(* CODESYS project CodeSys_main.project (continued)
  5ce3da45-db07-42e7-a21c-a00fff4ed8f6|C:\Users\ggb\Documents\#PROJECTS\2016_06_29_Denmark\Visu\RightArrow_Bold.png
  5ce3da45-db07-42e7-a21c-a00fff4ed8f6|C:\Users\ggb\Documents\#PROJECTS\2016_06_29_Denmark\Visu\Parameters_0.png
  5ce3da45-db07-42e7-a21c-a00fff4ed8f6|C:\Users\ggb\Documents\#PROJECTS\2016_06_29_Denmark\Pictures\071-060_Kameraprüfen.jpg
  5ce3da45-db07-42e7-a21c-a00fff4ed8f6|C:\Users\ggb\Documents\#PROJECTS\2016_06_29_Denmark\Visu\Manual_0.png
  5ce3da45-db07-42e7-a21c-a00fff4ed8f6|C:\Users\ggb\Documents\#PROJECTS\2016_06_29_Denmark\Pictures\071-046b_Magazin.jpg
  5ce3da45-db07-42e7-a21c-a00fff4ed8f6|C:\Users\ggb\Documents\#PROJECTS\2016_06_29_Denmark\Pictures\071-050a_Bohren EA.jpg
  5ce3da45-db07-42e7-a21c-a00fff4ed8f6|C:\Users\ggb\Documents\#PROJECTS\2016_06_29_Denmark\Visu\RightArrow_Bold.png
  5ce3da45-db07-42e7-a21c-a00fff4ed8f6|C:\Users\ggb\Documents\#PROJECTS\2016_06_29_Denmark\Visu\Manual_1.png
  5ce3da45-db07-42e7-a21c-a00fff4ed8f6|C:\Users\ggb\Documents\#PROJECTS\2016_06_29_Denmark\Visu\Plus.png
  5ce3da45-db07-42e7-a21c-a00fff4ed8f6|C:\Users\ggb\Documents\#PROJECTS\2016_06_29_Denmark\Visu\LeftArrow_Bold.png
  5ce3da45-db07-42e7-a21c-a00fff4ed8f6|C:\Users\ggb\Documents\#PROJECTS\2016_06_29_Denmark\Visu\German.gif
  5ce3da45-db07-42e7-a21c-a00fff4ed8f6|C:\Users\ggb\Documents\#PROJECTS\2016_06_29_Denmark\Pictures\071-030_Modul Trocknen.jpg
  5ce3da45-db07-42e7-a21c-a00fff4ed8f6|C:\Users\ggb\Documents\#PROJECTS\2016_06_29_Denmark\Visu\CheckBox_1.png
  5ce3da45-db07-42e7-a21c-a00fff4ed8f6|C:\Users\ggb\Documents\#PROJECTS\2016_06_29_Denmark\Visu\Manual_1.png
  5ce3da45-db07-42e7-a21c-a00fff4ed8f6|C:\Users\ggb\Documents\#PROJECTS\2016_06_29_Denmark\Visu\RightArrow.png
  5ce3da45-db07-42e7-a21c-a00fff4ed8f6|C:\Users\ggb\Documents\#PROJECTS\2016_06_29_Denmark\Visu\English.gif
  5ce3da45-db07-42e7-a21c-a00fff4ed8f6|C:\Users\ggb\Documents\#PROJECTS\2016_06_29_Denmark\Pictures\cpFactory_Conveyor.png
  5ce3da45-db07-42e7-a21c-a00fff4ed8f6|C:\Users\ggb\Documents\#PROJECTS\2016_06_29_Denmark\Visu\Parameters_0.png
  5ce3da45-db07-42e7-a21c-a00fff4ed8f6|C:\Users\ggb\Documents\#PROJECTS\2016_06_29_Denmark\Visu\Stopper.jpg
  5ce3da45-db07-42e7-a21c-a00fff4ed8f6|C:\Users\ggb\Documents\#PROJECTS\2016_06_29_Denmark\Visu\RightArrow_Bold.png
  5ce3da45-db07-42e7-a21c-a00fff4ed8f6|C:\Users\ggb\Documents\#PROJECTS\2016_06_29_Denmark\Visu\Home_1.png
  5ce3da45-db07-42e7-a21c-a00fff4ed8f6|C:\Users\ggb\Documents\#PROJECTS\2016_06_29_Denmark\Visu\CheckBox_0.png
  5ce3da45-db07-42e7-a21c-a00fff4ed8f6|C:\Users\ggb\Documents\#PROJECTS\2016_06_29_Denmark\Pictures\071-050a_Bohren EA.jpg
  5ce3da45-db07-42e7-a21c-a00fff4ed8f6|C:\Users\ggb\Documents\#PROJECTS\2016_06_29_Denmark\Visu\German.gif
  5ce3da45-db07-42e7-a21c-a00fff4ed8f6|C:\Users\ggb\Documents\#PROJECTS\2016_06_29_Denmark\Visu\English.gif
  5ce3da45-db07-42e7-a21c-a00fff4ed8f6|C:\Users\ggb\Documents\#PROJECTS\2016_06_29_Denmark\Visu\Plus.png
  5ce3da45-db07-42e7-a21c-a00fff4ed8f6|C:\Users\ggb\Documents\#PROJECTS\2016_06_29_Denmark\Visu\Parameters_1.png
*)

// Data Types/HMI and SCADA/st_WinCC
/////////////////////////////////
/////////////////////////////////
TYPE st_WinCC :
STRUCT
	/// activate Automatic mode
	xAuto: BOOL;
	/// activate Reset mode
	xReset: BOOL;
	/// Stop at cycle end
	xCycleEnd: BOOL;
	/// activate Manual mode
	xManual: BOOL;
	/// activate Teach mode
	xTeach: BOOL;
	/// Quit Error from WinCC
	xQuit: BOOL;
	/// Clear RFID Data (without CarrierID)
	xClrRFID: BOOL;
END_STRUCT
END_TYPE

// Data Types/SAP/sub_structures/st_Par_Req

TYPE st_Par_Req :
STRUCT
	sSfc		: STRING(18);
	sDcGroup	: STRING(12);
	sName1		: STRING(30);
	iValue1		: INT;
	sName2		: STRING(30);
	iValue2		: INT;
	sName3		: STRING(30);
	iValue3		: INT;
	sName4		: STRING(30);
	iValue4		: INT;
	iCamResult	: INT;
END_STRUCT
END_TYPE

// Data Types/Error/st_InteractiveError
//////////////////////////////////////////////
//////////////////////////////////////////////
TYPE st_InteractiveError :
STRUCT
	/// Interactive error is active
	xError: BOOL;
	/// Message ID (ID of the InteractiveErrors textlist row)
	sMessageID: STRING;
	/// The actual state of the stopper
	uiState: UINT;
	/// The state of stopper after pushing the Ignore button
	uiIgnoreState: UINT;
	/// The state of stopper after pushing the Abort button
	uiAbortState: UINT;
	/// Repeat button was pushed
	xBtnRepeat: BOOL;
	/// Ignore button was pushed
	xBtnIgnore: BOOL;
	/// Abort button was pushed
	xBtnAbort: BOOL;
	// Reject order button was pushed
	xBtnRejectOrder: BOOL;
END_STRUCT
END_TYPE

// Data Types/HMI and SCADA/CDPX/st_StopperSensorSignals
TYPE st_StopperSensorSignals :
STRUCT
	xInductive_1		: BOOL;
	xInductive_2		: BOOL;
	xInductive_3		: BOOL;
	xInductive_4		: BOOL;
	xStpDownSensor		: BOOL;
	xStpDownOutpu		: BOOL;
	sInductive_1		: STRING(5);
	sInductive_2		: STRING(5);
	sInductive_3		: STRING(5);
	sInductive_4		: STRING(5);
	sStpDownSensor		: STRING(5);
	sStpDownOutpu		: STRING(5);
	sRfid				: STRING(5);
	xTagPresent			: BOOL;
	xReady				: BOOL;
	xBusy				: BOOL;
	xError				: BOOL;
	xTimeOut			: BOOL;		
END_STRUCT
END_TYPE

// Data Types/HMI and SCADA/st_ManualWorkplace
TYPE st_ManualWorkplace :
STRUCT
	sURL				: STRING;
	xManualJob			: BOOL;
	xManualJobStarted	: BOOL;
	xManualJobFinished	: BOOL;
	xManualJobCanceled	: BOOL;
END_STRUCT
END_TYPE

// Data Types/HMI and SCADA/CDPX/st_InterctiveErrors
TYPE st_InterctiveErrors :
STRUCT
	xIntDefault		: BOOL;
	xIntMES			: BOOL;
	xIntSAP			: BOOL;
	xIntApp			: BOOL;
	xIntMan			: BOOL;
	xIntKuka		: BOOL;
	
	sURL			: STRING;
	uiIntMsgID		: UINT;
	uiIntState		: UINT;
	uiIntIgnore		: UINT;
	uiIntAbort		: UINT;
	uiSapOp			: UDINT;
	uiSapPos		: UDINT;
	sSapError		: STRING;
	udiSapSfc		: UDINT;	
END_STRUCT
END_TYPE

// Data Types/HMI and SCADA/CDPX/st_Errors
TYPE st_Errors :
STRUCT
	xError			: BOOL;
	uiLevel			: UINT;
	uiMsgNum		: UINT;
	sErrorID		: STRING[4);
	sDateTime		: STRING;
END_STRUCT
END_TYPE

// Data Types/Error/st_RobotError
TYPE st_RobotError :
STRUCT
	/// Interactive error is active
	xError: BOOL;
	/// Message ID (ID of the InteractiveErrors textlist row)
	sMessageID: STRING;
	/// The state of stopper after pushing the Retry button
	uiRetryState: UINT;
	/// The state of stopper after pushing the Exit button
	uiExitState: UINT;
	/// Retry button was pushed
	xBtnRetry: BOOL;
	/// Exit button was pushed
	xBtnExit: BOOL;
END_STRUCT
END_TYPE

// Data Types/Application/st_AppControl
TYPE st_AppControl :
STRUCT
	xStart		: BOOL;
	xReset		: BOOL;
	xStop		: BOOL;
	uiOpNo		: UINT;
	auiPar		: ARRAY [0..3] OF UINT;
	udiONo		: UDINT;
	uiOPos		: UINT;
END_STRUCT
END_TYPE

// Data Types/HMI and SCADA/CDPX/st_ConveyorSignals
TYPE st_ConveyorSignals :
STRUCT
	xConvMovingLeft		: BOOL;
	xConvMovingRight	: BOOL;
	xConvMovingSlow		: BOOL;
	
	sConvLeft			: STRING(5);
	sConvRight			: STRING(5);
	sConvSlow			: STRING(5);	
END_STRUCT
END_TYPE

// Data Types/Error/u_Error
////////////////////////////////////////////////////////////////////////////////////////
/////////////////////////////////////////////////////////////////////////////////////////
TYPE u_Error :

UNION
	/// Long Word (64 bit) for error bits
	lwError: LWORD;
	/// 4 times Word for WinCC visualization
	stErrorWords: st_ErrorWords;
END_UNION

END_TYPE

// Data Types/Error/st_Error
///////////////////////////////////
///////////////////////////////////
TYPE st_Error :
STRUCT
	/// Union to store Level 0 errors in LWORD and 4xWORD for WinCC
	uL0: u_Error;
	/// Union to store Level 1 errors in LWORD and 4xWORD for WinCC
	uL1: u_Error;
	/// Union to store Level 2 errors in LWORD and 4xWORD for WinCC	
	uL2: u_Error;
	/// Error flags
	xSF0: BOOL;
	/// summary error flag Level 1
	xSF1: BOOL;
	/// summary error flag Level 2
	xSF2: BOOL;
	/// global error flag (SF0 or SF1)
	xSF: BOOL;
	/// extended (100ms) global error flag
	xSF_ext: BOOL;
	/// confirm error
	xQuit: BOOL;
END_STRUCT
END_TYPE

// Data Types/SAP/sub_structures/st_Start_Req

TYPE st_Start_Req :
STRUCT
	sSfc	: STRING(18);
	sItem	: STRING(18);
END_STRUCT
END_TYPE

// Data Types/SAP/st_CompleteSfc

TYPE st_CompleteSfc :
STRUCT
	Req		: st_Comp_Req;
	Res		: st_Comp_Res;
	Com		: st_Com;
END_STRUCT
END_TYPE

// Data Types/HMI and SCADA/st_ButtonState
TYPE st_ButtonState :
STRUCT
	xPressed	: BOOL;
	xActive		: BOOL;
	xDisabled	: BOOL;
END_STRUCT
END_TYPE

// Data Types/SAP/st_ParametricData

TYPE st_ParametricData :
STRUCT
	Req		: st_Par_Req;
	Com		: st_Com;
END_STRUCT
END_TYPE

// Data Types/Application/st_AppSettings
TYPE st_AppSettings :
STRUCT
	xActive			: BOOL := TRUE;
	xStopBelt		: BOOL;
	xCarrierInit	: BOOL;
	uiCarrierInitNum: UINT := 1;
END_STRUCT
END_TYPE

// Data Types/HMI and SCADA/CDPX/st_AppButtonControl
TYPE st_AppButtonControl :
STRUCT
	xButton		: BOOL;
	sButton		: STRING(16);	
END_STRUCT
END_TYPE

// Data Types/SAP/sub_structures/st_Com

TYPE st_Com :
STRUCT
	iTrigger		: INT;
	iResponse		: INT;
	bError			: BIT;
	sError			: STRING(128);
END_STRUCT
END_TYPE

// Data Types/Application/st_AppState
TYPE st_AppState :
STRUCT
	xReady					: BOOL;
	xError					: BOOL;
	xInitPos				: BOOL;
	uiReturnCode			: UINT;
END_STRUCT
END_TYPE

// Data Types/HMI and SCADA/CDPX/st_StopperButtonState
TYPE st_StopperButtonState :
STRUCT
	xInit		: BOOL;
	xRead		: BOOL;
	xWrite		: BOOL;
	xDeleteData	: BOOL;
	xStpMveDown	: BOOL;
	xStpMveUp	: BOOL;
END_STRUCT
END_TYPE

// Data Types/Error/st_ErrorWords
/////////////////////////
/////////////////////////
TYPE st_ErrorWords :
STRUCT
	wErrorWord0: WORD;
	wErrorWord1: WORD;
	wErrorWord2: WORD;
	wErrorWord3: WORD;
END_STRUCT
END_TYPE

// Data Types/SAP/sub_structures/st_Start_Res

TYPE st_Start_Res :
STRUCT
	sDcGroup	: STRING(12);
	sName1		: STRING(30);
	iValue1		: INT;
	sName2		: STRING(30);
	iValue2		: INT;
	sName3		: STRING(30);
	iValue3		: INT;
	sName4		: STRING(30);
	iValue4		: INT;
	sItem		: STRING(18);
	sItemRev	: STRING(3);
	sSfc		: STRING(10);	
END_STRUCT
END_TYPE

// Data Types/HMI and SCADA/CDPX/st_CdpxButtonState
TYPE st_CdpxButtonState :
STRUCT
	xClearError		: BOOL;
	xOperationMode	: BOOL;
	xOverview     	: BOOL;
	xUser         	: BOOL;
	xHome         	: BOOL;
	xSetupMode    	: BOOL;
	xParameter    	: BOOL;
	xSystem       	: BOOL;
	xApp_1        	: BOOL;
	xApp_2        	: BOOL;
	xStp_1        	: BOOL;
	xStp_2        	: BOOL;
	xBelt         	: BOOL;
	xApp          	: BOOL;
	xTrans_1      	: BOOL;
	xTrans_2      	: BOOL;
	xSwLanguage		: BOOL;
	xCloseDialog	: BOOL;
END_STRUCT
END_TYPE

// Data Types/SAP/ManualWork/st_MesRcvData_ManualWork
TYPE st_MesRcvData_ManualWork :
STRUCT
	stHeader		: dc_ecp.st_MES4_QueryHeader;
	sOderDes		: STRING[60];
	sPartDes		: STRING[20];
END_STRUCT
END_TYPE

// Data Types/Application/st_AppInfo
TYPE st_AppInfo :
STRUCT
	auiOperations			: ARRAY [0..15] OF UINT;
	byNumberOfOperations	: BYTE;
END_STRUCT
END_TYPE

// Data Types/SAP/sub_structures/st_Comp_Req

TYPE st_Comp_Req :
STRUCT
	sSfc	: STRING(18);
END_STRUCT
END_TYPE

// Data Types/HMI and SCADA/CDPX/st_AppSensors
TYPE st_AppSensors :
STRUCT
	xSensor		: BOOL;
	sSensor		: STRING(16);
END_STRUCT
END_TYPE

// Data Types/SAP/sub_structures/st_Comp_Res

TYPE st_Comp_Res :
STRUCT
	sOp		: STRING(4);
	sOpRev	: STRING(3);
END_STRUCT
END_TYPE

// Data Types/st_GetShuntId
TYPE st_GetShuntId :
STRUCT
	uiSourceId			: UINT;
	uiSourcePosition	: UINT;
	uiTargetId			: UINT;
	uiTargetPosition	: UINT;
END_STRUCT
END_TYPE

// Data Types/Error/st_ErrorEvent
///////////////////////////////////
///////////////////////////////////
TYPE st_ErrorEvent :
STRUCT
	/// Error ID (ID of the Errors textlist row)
	sErrorID: STRING := 'No error';
	/// Text message (It does not contains anyting, it is only to show an additional column in the visualization)
	sErrorText: STRING;
	/// String of the date and time
	sDateTime: STRING;
END_STRUCT
END_TYPE

// Data Types/HMI and SCADA/st_TransitionData
TYPE st_TransitionData :
STRUCT
	uiCondIn	: UINT;
	uiPar1		: UINT;
	uiPar2		: UINT;
	uiPar3		: UINT;
	uiPar4		: UINT;
	xAppEn		: BOOL;
	uiCondOut	: UINT;
	uiCondAbort	: UINT;
	byStopper	: BYTE;
END_STRUCT
END_TYPE

// Data Types/SAP/st_StartSfc

TYPE st_StartSfc :
STRUCT
	Req	: st_Start_Req;
	Res	: st_Start_Res;
	Com	: st_Com;
END_STRUCT
END_TYPE

// Data Types/HMI and SCADA/CDPX/st_ConveyorButtonState
TYPE st_ConveyorButtonState :
STRUCT
	xConvLeft		: BOOL;
	xConvRight		: BOOL;
	xConvSlow		: BOOL;
END_STRUCT
END_TYPE

// Global Variables/fromCDPX
{attribute 'qualified_only'}
VAR_GLOBAL
	uiMode									: UINT;
	uiDummy									: UINT;
	stCdpxButtonState						: st_CdpxButtonState;
	
	
	stHome_OperationMode_Reset		 		: st_ButtonState;
	stHome_OperationMode_Automatic		 	: st_ButtonState;
	stHome_OperationMode_Setup 				: st_ButtonState;
	stHome_OperationMode_CycleEnd 			: st_ButtonState;
	
	stSetupMode_Stopper1_Init		 		: st_ButtonState;
	stSetupMode_Stopper1_Read			 	: st_ButtonState;
	stSetupMode_Stopper1_Write 				: st_ButtonState;
	stSetupMode_Stopper1_DeleteData 		: st_ButtonState;

	stSetupMode_Stopper2_Init		 		: st_ButtonState;
	stSetupMode_Stopper2_Read			 	: st_ButtonState;
	stSetupMode_Stopper2_Write 				: st_ButtonState;
	stSetupMode_Stopper2_DeleteData 		: st_ButtonState;
	
	stInteractiveMessage_Repeat 			: st_ButtonState;
	stInteractiveMessage_Ignore	 			: st_ButtonState;
	stInteractiveMessage_Abort				: st_ButtonState;	
	stInteractiveMessage_RejectOrder		: st_ButtonState;	
	
	stManualWorkplace						: st_ManualWorkplace;
	stRobotError							: st_RobotError;	
	astStopperButton						: ARRAY [0..1] OF st_StopperButtonState;
	astAppSetting							: ARRAY [0..1] OF st_AppSettings;
	astAppButtonControl						: ARRAY [0..15] OF st_AppButtonControl;
	astTransitionTable_1					: ARRAY [0..10] OF st_TransitionData;
	astTransitionTable_2					: ARRAY [0..10] OF st_TransitionData;	
	astConveyorButtonState					: ARRAY [0..2] OF st_ConveyorButtonState; 
END_VAR

// APP_FILLING/Application/IO
//{attribute 'qualified_only'} - removed to access variables without "DigitalIO." 
VAR_GLOBAL
	// Application Type Identifier
	xAppID AT %QX0.7: BOOL := TRUE;
	// Push Piston forward
	xPistonOn AT %QX0.0: BOOL := FALSE;
	// Turns pump on
	xPumpOn AT %QX0.2: BOOL := FALSE;
	// Indicates if the app is powered on or off
	xIsOn AT %QX0.6: BOOL := TRUE;
	// Indicates which module (09 or 08) the app is mounted on
	xModuleID AT %IX0.7: BOOL;
END_VAR

// Global Variables/Standards
VAR_GLOBAL
	/// First-Cycle-Flag
	xFirstCycle: BOOL := TRUE;
	/// Initialization flag
	xInit: BOOL;
	/// Station is in Initial Position
	xInitPos: BOOL;
	/// Startup like warmstart
	xSoftReset: BOOL;
	/// Application program is idle	
	xAppIdle: BOOL;
	/// Application program is busy
	xAppBusy: BOOL;
	/// Automatic Mode is active
	xAuto: BOOL;
	/// Automatic Start is enable
	xAutoEn: BOOL;
	/// Reset Mode is active
	xReset: BOOL;
	/// Reset Start is enable
	xResetEn: BOOL;
	/// Reset sequence is finished
	xResetRdy: BOOL;
	/// Manual Mode is active
	xManual: BOOL;
	/// Manual Start is enable
	xManualEn: BOOL;
	/// Teach Mode is active	
	xTeach: BOOL;
	/// Teach Start is enable
	xTeachEn: BOOL;
	/// Stop at cycle end is active	
	xCycleEnd: BOOL;
	/// Stop at cycle end is enable
	xCycleEndEn: BOOL;
	/// Reset Automatic Start flag
	xAutoReset: BOOL := FALSE;
	/// Stopper ST1 in idle state          		
	xSt1_Idle: BOOL;
	/// Stopper ST2 in idle state          		
	xSt2_Idle: BOOL;
	/// Stopper ST2 in idle state          		
	xSt3_Idle: BOOL;
	/// Resource is busy
	xBusy: BOOL;
	/// MES mode is active
	xMES: BOOL;
	/// SAP mode is active
	xSAP: BOOL;
	/// Struct with 64 Error Flags
	stError: st_Error;
	/// Structure with WinCC variables     
	stWinCC: st_WinCC;
	/// Structure with HMI variables
	stHMI: st_WinCC;
	//Semaphore for gate
	xSema : BOOL;
	// Semaphore for shunt
	xSemaShunt	: BOOL;
END_VAR

// Global Variables/toCDPX
{attribute 'qualified_only'}
VAR_GLOBAL
	sModule						: STRING(32);
	byOpMode					: BYTE;
	byScreenTitle				: BYTE;
	xManual						: BOOL;
	xAuto						: BOOL;
	xSAP						: BOOL;
	xMES						: BOOL;
	xDefault					: BOOL;
	auiCarrierInitNum			: ARRAY [0..1] OF UINT;
	uiNumOfApplications			: UINT;
	uiNumOfStoppers				: UINT;
	uiNumOfBelts				: UINT;
	auiCondIn					: ARRAY [0..1] OF UINT;
	auiCondOut					: ARRAY [0..1] OF UINT;
	sTime						: STRING;
	sDate						: STRING;
	stInteractiveErrors			: st_InterctiveErrors;
	astErrors					: ARRAY [1..20] OF st_Errors;
	astRfidData					: ARRAY [0..1] OF dc_ecp.st_CPF_VisuData;
	astSensorSignals			: ARRAY [0..1] OF st_StopperSensorSignals;
	astConveyorSignals			: ARRAY [0..2] OF st_ConveyorSignals;
	astAppState					: ARRAY [0..1] OF st_AppState;
	astAppControl				: ARRAY [0..1] OF st_AppControl;	
	astAppSensors				: ARRAY [0..31] OF st_AppSensors;
	auiValues					: ARRAY [0..31] OF UINT;	
	astAppControlONo: UDINT := 0;
END_VAR

// Global Variables/SAP
{attribute 'qualified_only'}
VAR_GLOBAL
	Start			: st_StartSfc;
	Par				: st_ParametricData;
	Comp			: st_CompleteSfc;
END_VAR

// Global Variables/SAPInit
{attribute 'qualified_only'}
VAR_GLOBAL
	Start			: st_StartSfc;
	Par				: st_ParametricData;
	Comp			: st_CompleteSfc;
END_VAR

// Global Variables/SAPHMI
{attribute 'qualified_only'}
VAR_GLOBAL
	uiOp		: UDINT;
	uiPos		: UDINT;
	sError		: STRING;
	udiSfc		: UDINT;	
END_VAR

// MODULE_PLC09/Application/Variables/IO
VAR_GLOBAL
	

	///////////////////////////
	// Inputs
	///////////////////////////
	
	xBG20		AT %IX1.0	: BOOL;	// Stopper released
	xBG21		AT %IX1.1	: BOOL;	// Carrier available
	xBG22		AT %IX1.2	: BOOL;	// Carrier ID bit 0
	xBG23		AT %IX1.3	: BOOL;	// Carrier ID bit 1
	xBG24		AT %IX1.4	: BOOL;	// Carrier ID bit 2
	xEmg		AT %IX0.0	: BOOL;	// Emergency stop
	
	///////////////////////////
	// Outputs
	///////////////////////////	
	
	xMB20		AT %QX1.0	: BOOL;	// Release stopper
	xQA1_LEFT	AT %QX0.5	: BOOL;	// Conveyor to the left
	xQA1_RIGHT	AT %QX0.4	: BOOL;	// Conveyor to the right
	xQA1_SLOW	AT %QX0.6	: BOOL;	// Conveyor Slow
	xQA1_STOP	AT %QX0.7	: BOOL;	// Conveyor Stop
	// Application Identifier
	xAPP_ID AT %IX0.1: BOOL;
	
	
	
	
	// Application power status
	xAppIsOn AT %IX0.2: BOOL;
	// Module Identifier Bit
	xModuleID AT %QX0.0: BOOL := FALSE;
END_VAR

// MODULE_PLC09/Application/Variables/NVL_PLC09_REC_FILLING
//This gobal variable list is received via the network.
//Sender: NVL_FILLING_SEND [APP_FILLING: PLC Logic: Application]
//Protocol: UDP

VAR_GLOBAL
	isDone: BOOL := FALSE;
	isOn: BOOL := FALSE;
END_VAR

// MODULE_PLC09/Application/Variables/NVL_PLC09_SEND
VAR_GLOBAL
	Ready: BOOL := FALSE;
END_VAR

// MODULE_PLC08/Application/Variables/IO
VAR_GLOBAL
	

	///////////////////////////
	// Inputs
	///////////////////////////
	
	xBG20		AT %IX1.0	: BOOL;	// Stopper released
	xBG21		AT %IX1.1	: BOOL;	// Carrier available
	xBG22		AT %IX1.2	: BOOL;	// Carrier ID bit 0
	xBG23		AT %IX1.3	: BOOL;	// Carrier ID bit 1
	xBG24		AT %IX1.4	: BOOL;	// Carrier ID bit 2
	xEmg		AT %IX0.0	: BOOL;	// Emergency stop
	
	///////////////////////////
	// Outputs
	///////////////////////////	
	
	xMB20		AT %QX1.0	: BOOL;	// Release stopper
	xQA1_LEFT	AT %QX0.5	: BOOL;	// Conveyor to the left
	xQA1_RIGHT	AT %QX0.4	: BOOL;	// Conveyor to the right
	xQA1_SLOW	AT %QX0.6	: BOOL;	// Conveyor Slow
	xQA1_STOP	AT %QX0.7	: BOOL;	// Conveyor Stop
	// Application Identifier
	xAPP_ID AT %IX0.1: BOOL;
	
	
	// Application power status
	xAppIsOn AT %IX0.2: BOOL;
	// Module Identifier Bit
	xModuleID AT %QX0.0: BOOL := TRUE;
END_VAR

// MODULE_PLC08/Application/Variables/NVL_PLC08_SEND
VAR_GLOBAL
	Ready: BOOL := FALSE;
END_VAR

// APP_FILLING/Application/NVL_FILLING_SEND
VAR_GLOBAL
	isDone: BOOL := FALSE;
	isOn: BOOL := FALSE;
END_VAR

// APP_FILLING/Application/NVL_FILLING_REC_09
//This gobal variable list is received via the network.
//Sender: NVL_PLC09_SEND [MODULE_PLC09: PLC Logic: Application]
//Protocol: UDP

VAR_GLOBAL
	Ready: BOOL := FALSE;
END_VAR

// APP_STOPPERING/Application/IO
//{attribute 'qualified_only'} - removed to access variables without "DigitalIO." 
VAR_GLOBAL
	// Application Type Identifier
	xAppID AT %QX0.7: BOOL := FALSE;
	// Push Piston forward
	xPistonOn AT %QX0.0: BOOL := FALSE;
	// Pushes stoppering down to the containers
	xStopperingOn AT %QX0.2: BOOL := FALSE;
	// Indicates if the app is powered on or off
	xIsOn AT %QX0.6: BOOL := TRUE;
	// Indicates which module (09 or 08) the app is mounted on
	xModuleID AT %IX0.7: BOOL;
END_VAR

// APP_STOPPERING/Application/NVL_STOPPERING_SEND
VAR_GLOBAL
	isDone: BOOL := FALSE;
END_VAR

// APP_STOPPERING/Application/NVL_STOPPERING_REC_08
//This gobal variable list is received via the network.
//Sender: NVL_PLC08_SEND [MODULE_PLC08: PLC Logic: Application]
//Protocol: UDP

VAR_GLOBAL
	Ready: BOOL := FALSE;
END_VAR

// MODULE_PLC08/Application/Variables/NVL_PLC08_REC_STOPPERING
//This gobal variable list is received via the network.
//Sender: NVL_STOPPERING_SEND [APP_STOPPERING: PLC Logic: Application]
//Protocol: UDP

VAR_GLOBAL
	isDone: BOOL := FALSE;
END_VAR

// MODULE_PLC08/Application/Variables/NVL_PLC08_REC_FILLING
//This gobal variable list is received via the network.
//Sender: NVL_FILLING_SEND [APP_FILLING: PLC Logic: Application]
//Protocol: UDP

VAR_GLOBAL
	isDone: BOOL := FALSE;
	isOn: BOOL := FALSE;
END_VAR

// APP_STOPPERING/Application/NVL_STOPPERING_REC_09
//This gobal variable list is received via the network.
//Sender: NVL_PLC09_SEND [MODULE_PLC09: PLC Logic: Application]
//Protocol: UDP

VAR_GLOBAL
	Ready: BOOL := FALSE;
END_VAR

// APP_FILLING/Application/NVL_FILLING_REC_08
//This gobal variable list is received via the network.
//Sender: NVL_PLC08_SEND [MODULE_PLC08: PLC Logic: Application]
//Protocol: UDP

VAR_GLOBAL
	Ready: BOOL := FALSE;
END_VAR

// MODULE_PLC09/Application/Variables/NVL_PLC09_REC_STOPPERING
//This gobal variable list is received via the network.
//Sender: NVL_STOPPERING_SEND [APP_STOPPERING: PLC Logic: Application]
//Protocol: UDP

VAR_GLOBAL
	isDone: BOOL := FALSE;
END_VAR

// MODULE_PLC09/Application/Programs/MODULE_PLC09_MAIN
PROGRAM  MODULE_PLC09_MAIN
VAR
	state: UINT := 0;
	PLCid: STRING;
	RFID: dc_ecp.Dtm425;
	RfidData: dc_ecp.st_CPF_RfidData;
	ConveyorRight: BOOL;
	CarrierID: UINT := 0;
	TIMER: TON;
	WaitTime: TIME;
	AppType: STRING;
	PistonState: STRING := 'retracted';
	ServerCommand: STRING := 'wait';
	AppState: STRING := 'waiting';
	CarrierIdString: STRING := '0';
END_VAR

CASE state OF
	
	0: // init
	IO.xMB20 := FALSE; // raise stoppper
	RFID.ClearError();
	PLCid := 'STPLC_09';
	state := 5;
	
	5: // identify
	AppState := 'N/A';
	IF IO.xAppIsOn THEN
		IF IO.xAPP_ID THEN
			AppType := 'filling';
		ELSE
			AppType := 'stoppering';
		END_IF
		state:=10;
	END_IF
	
	10: // wait for RFID to clear
	AppState := 'starting';
	IF RFID.xReady THEN
		RFID.Connect(32, 0, 1);
		state:=20;
	END_IF
	
	20: // wait for RFID be ready then move conveyor
	//CarrierID := 0;
	IF RFID.xReady AND IO.xAppIsOn THEN
		AppState := 'ready';
		IF ServerCommand = 'begin' THEN
			AppState := 'waiting';
			IO.xMB20 := TRUE;
			IO.xQA1_RIGHT := TRUE; // Move conveyor right
			state:=30;
		END_IF
	ELSE
		AppState := 'N/A';
	END_IF
	
	30: // wait for carrier to be available
	IF IO.xBG21 THEN
		IO.xQA1_RIGHT := FALSE; // stop conveyor
		IO.xMB20 := FALSE; // lower stoppper
		state:=40;
	END_IF
	
	
	40: // wait for RFID to read then send
	IF RFID.xReady THEN
		RFID.ReadTag(uiStartAddress := 0, uiDataLength := SIZEOF(RfidData), ADR(RfidData));
		state := 42;
	END_IF
	
	42:
	IF RFID.xReady THEN
		CarrierID := dc_ecp.SwapWord(RfidData.uiCarrierID); // swap bit order
		
		IF CarrierID > 0 THEN
			AppState := 'ready';
			state := 45;
		ELSE
			AppState := 'waiting';
		END_IF
	END_IF
	
	45: // wait for server to tell if pass or go
	IF ServerCommand = 'valid' THEN
		IF AppType = 'filling' THEN
			AppState := 'filling';
			state := 46;
		ELSIF AppType = 'stoppering' THEN
			AppState := 'stoppering';
			state := 46;
		END_IF
	ELSIF ServerCommand = 'pass' THEN
		AppState := 'passing';
		state := 100;
	END_IF
	
	46:
	NVL_PLC09_SEND.Ready := TRUE;
	WaitTime := STRING_TO_TIME('T#500ms');
	TIMER(IN := TRUE, PT := WaitTime);
	IF TIMER.Q = TRUE THEN 
		TIMER(IN := FALSE);
		NVL_PLC09_SEND.Ready := FALSE;
		state := 50;
	END_IF
	
	
	50: // wait for task to complete, then report back
	IF AppType = 'stoppering' THEN
		IF NVL_PLC09_REC_STOPPERING.isDone THEN
			AppState := 'done';
			state := 55;
		END_IF
	ELSIF AppType = 'filling' THEN
		IF NVL_PLC09_REC_FILLING.isDone THEN
			AppState := 'done';
			state := 55;
		END_IF
	END_IF
	
	55: // wait for server to tell it to move on
	IF ServerCommand = 'transfer' THEN
		state := 100;
	END_IF
	

	
	100: // pass move conveyor again, give 1 sec breathing room
	IO.xMB20 := TRUE; // release stopper
	IF IO.xBG20 THEN // checks if stopper has been released
		IO.xQA1_RIGHT := TRUE; // move conveyor right
		WaitTime := STRING_TO_TIME('T#2000ms');
		timer(IN:=TRUE,PT:=WaitTime);
		state := 105;
	END_IF
	
	105: // wait for timer then restart
	IF timer.Q = TRUE THEN
		timer(IN:=FALSE);
		IF ServerCommand = 'pass' THEN
			AppState := 'passed';
		ELSIF ServerCommand = 'transfer' THEN
			AppState := 'done';
		END_IF
		state := 30;
		CarrierID := 0;
		ServerCommand := 'begin';
	END_IF
	
	
	
END_CASE
RFID();
timer();

END_PROGRAM

// APP_FILLING/Application/APP_FILLING_MAIN
PROGRAM APP_FILLING_MAIN
VAR
	state: UINT := 0;
	APPid: STRING;
	TIMER: TON;
	WaitTime: TIME;
	ModuleID: STRING;
END_VAR

CASE state OF
	
	0: // init
	APPid := 'APP_FILLINGs';
	IO.xPistonOn := FALSE;
	IO.xPumpOn := FALSE;
	IO.xIsOn := TRUE;
	IO.xAppID := TRUE;
	NVL_FILLING_SEND.isOn := TRUE;
	state := 10;
	
	10: //  Read Module id
	IF IO.xModuleID = TRUE THEN
		ModuleID := '08';
	ELSIF IO.xModuleID = FALSE THEN
		ModuleID := '09';
	END_IF
	state := 15;
	
	15: // wait for module to be ready
	IF ModuleID = '08' THEN
		IF NVL_FILLING_REC_08.Ready THEN
			NVL_FILLING_SEND.isDone := FALSE;
			state := 20;
		END_IF
	ELSIF ModuleID = '09' THEN
		IF NVL_FILLING_REC_09.Ready THEN
			NVL_FILLING_SEND.isDone := FALSE;
			state := 20;
		END_IF
	END_IF
	
	20: // Push piston forward and wait 5 sec
	IO.xPistonOn := TRUE;
	WaitTime := STRING_TO_TIME ('T#500ms'); // Converts text string to time value --> WaitTime is then 5 sec
	TIMER(IN := TRUE, PT := WaitTime); // Activates the timer and the timers preset time --> The time where the piston is active
	IF Timer.Q = TRUE THEN 
		TIMER(IN := FALSE);
		state := 25;
	END_IF
	
	25: // activate pump for 200ms
	//IO.PistonOn := FALSE;
	IO.xPumpOn := TRUE;
	WaitTime := STRING_TO_TIME ('T#200ms'); // Converts text string to time value --> WaitTime is then 5 sec
	TIMER(IN := TRUE, PT := WaitTime); // Activates the timer and the timers preset time --> The time where the piston is active
	IF Timer.Q = TRUE THEN 
		TIMER(IN := FALSE);
		IO.xPumpOn := FALSE;
		state := 30;
	END_IF
	
	30: // Push piston backwards
	WaitTime := STRING_TO_TIME('T#500ms');
	TIMER(IN := TRUE, PT := WaitTime);
	IF TIMER.Q = TRUE THEN 
		TIMER(IN := FALSE);
		IO.xPistonOn := FALSE;
		state := 40;
	END_IF
	
	40: // Restart conveyor belts
	NVL_FILLING_SEND.isDone := TRUE;
	WaitTime := STRING_TO_TIME('T#1000ms');
	TIMER(IN := TRUE, PT := WaitTime);
	IF TIMER.Q = TRUE THEN 
		TIMER(IN := FALSE);
		state := 15;
	END_IF
	
END_CASE

TIMER();

END_PROGRAM

// MODULE_PLC08/Application/Programs/MODULE_PLC08_MAIN
PROGRAM  MODULE_PLC08_MAIN
VAR
	state: UINT := 0;
	PLCid: STRING;
	RFID: dc_ecp.Dtm425;
	RfidData: dc_ecp.st_CPF_RfidData;
	ConveyorRight: BOOL;
	CarrierID: UINT := 0;
	TIMER: TON;
	WaitTime: TIME;
	AppType: STRING;
	PistonState: STRING := 'retracted';
	ServerCommand: STRING := 'wait';
	AppState: STRING := 'waiting';
END_VAR

CASE state OF
	
	0: // init
	IO.xMB20 := FALSE; // raise stoppper
	RFID.ClearError();
	PLCid := 'STPLC_08';
	state := 5;
	
	5: // identify
	AppState := 'N/A';
	IF IO.xAppIsOn THEN
		IF IO.xAPP_ID THEN
			AppType := 'filling';
		ELSE
			AppType := 'stoppering';
		END_IF
		state:=10;
	END_IF
	
	10: // wait for RFID to clear
	AppState := 'starting';
	IF RFID.xReady THEN
		RFID.Connect(32, 0, 1);
		state:=20;
	END_IF
	
	20: // wait for RFID be ready then move conveyor
	//CarrierID := 0;
	IF RFID.xReady AND IO.xAppIsOn THEN
		AppState := 'ready';
		IF ServerCommand = 'begin' THEN
			AppState := 'waiting';
			IO.xMB20 := TRUE;
			IO.xQA1_RIGHT := TRUE; // Move conveyor right
			state:=30;
		END_IF
	ELSE
		AppState := 'N/A';
	END_IF
	
	30: // wait for carrier to be available
	IF IO.xBG21 THEN
		IO.xQA1_RIGHT := FALSE; // stop conveyor
		IO.xMB20 := FALSE; // lower stoppper
		state:=40;
	END_IF
	
	
	40: // wait for RFID to read then send
	IF RFID.xReady THEN
		RFID.ReadTag(uiStartAddress := 0, uiDataLength := SIZEOF(RfidData), ADR(RfidData));
		state := 42;
	END_IF
	
	42:
	IF RFID.xReady THEN
		CarrierID := dc_ecp.SwapWord(RfidData.uiCarrierID); // swap bit order
		
		IF CarrierID > 0 THEN
			AppState := 'ready';
			state := 45;
		ELSE
			AppState := 'waiting';
		END_IF
	END_IF
	
	45: // wait for server to tell if pass or go
	IF ServerCommand = 'valid' THEN
		IF AppType = 'filling' THEN
			AppState := 'filling';
			state := 46;
		ELSIF AppType = 'stoppering' THEN
			AppState := 'stoppering';
			state := 46;
		END_IF
	ELSIF ServerCommand = 'pass' THEN
		AppState := 'passing';
		state := 100;
	END_IF
	
	46: // tell app to start then wait
	NVL_PLC08_SEND.Ready := TRUE;
	WaitTime := STRING_TO_TIME('T#500ms');
	TIMER(IN := TRUE, PT := WaitTime);
	IF TIMER.Q = TRUE THEN 
		TIMER(IN := FALSE);
		NVL_PLC08_SEND.Ready := FALSE;
		state := 50;
	END_IF
	
	
	50: // wait for task to complete, then report back
	IF AppType = 'stoppering' THEN
		IF NVL_PLC08_REC_STOPPERING.isDone THEN
			AppState := 'done';
			state := 55;
		END_IF
	ELSIF AppType = 'filling' THEN
		IF NVL_PLC08_REC_FILLING.isDone THEN
			AppState := 'done';
			state := 55;
		END_IF
	END_IF
	
	55: // wait for server to tell it to move on
	IF ServerCommand = 'transfer' THEN
		state := 100;
	END_IF
	

	
	100: // pass move conveyor again, give 1 sec breathing room
	IO.xMB20 := TRUE; // release stopper
	IF IO.xBG20 THEN // checks if stopper has been released
		IO.xQA1_RIGHT := TRUE; // move conveyor right
		WaitTime := STRING_TO_TIME('T#2000ms');
		timer(IN:=TRUE,PT:=WaitTime);
		state := 105;
	END_IF
	
	105: // wait for timer then restart
	IF timer.Q = TRUE THEN
		timer(IN:=FALSE);
		IF ServerCommand = 'pass' THEN
			AppState := 'passed';
		ELSIF ServerCommand = 'transfer' THEN
			AppState := 'done';
		END_IF
		state := 20;
		CarrierID := 0;
		ServerCommand := 'begin';
	END_IF
	
	
	
END_CASE
RFID();
timer();

END_PROGRAM

// APP_STOPPERING/Application/APP_STOPPERING_MAIN
PROGRAM APP_STOPPERING_MAIN
VAR
	state: UINT := 0;
	APPid: STRING;
	TIMER: TON;
	WaitTime: TIME;
	ModuleID: STRING;
END_VAR

CASE state OF
	
	0: // init
	APPid := 'APP_STOPPERING';
	IO.xPistonOn := FALSE;
	IO.xIsOn := TRUE;
	IO.xAppID := FALSE;
	state := 10;
	
	10: // Read Module id
	IF IO.xModuleID = TRUE THEN
		ModuleID := '08';
	ELSIF IO.xModuleID = FALSE THEN
		ModuleID := '09';
	END_IF
	state := 15;
	
	15: // wait for module to be ready
	IF ModuleID = '08' THEN
		IF NVL_STOPPERING_REC_08.Ready THEN
			NVL_STOPPERING_SEND.isDone := FALSE;
			state := 20;
		END_IF
	ELSIF ModuleID = '09' THEN
		IF NVL_STOPPERING_REC_09.Ready THEN
			NVL_STOPPERING_SEND.isDone := FALSE;
			state := 20;
		END_IF
	END_IF
		
	
	20: // Push piston forward and wait 5 sec
	IO.xPistonOn := TRUE;
	WaitTime := STRING_TO_TIME ('T#500ms'); // Converts text string to time value --> WaitTime is then 5 sec
	TIMER(IN := TRUE, PT := WaitTime); // Activates the timer and the timers preset time --> The time where the piston is active
	IF Timer.Q = TRUE THEN 
		TIMER(IN := FALSE);
		state := 25;
	END_IF
	
	25: // activate stopper
	IO.xStopperingOn := TRUE;
	WaitTime := STRING_TO_TIME ('T#500ms'); // Converts text string to time value --> WaitTime is then 5 sec
	TIMER(IN := TRUE, PT := WaitTime); // Activates the timer and the timers preset time --> The time where the piston is active
	IF Timer.Q = TRUE THEN 
		TIMER(IN := FALSE);
		IO.xStopperingOn := FALSE;
		state := 30;
	END_IF
	
	30: // Push piston backwards
	WaitTime := STRING_TO_TIME('T#500ms');
	TIMER(IN := TRUE, PT := WaitTime);
	IF TIMER.Q = TRUE THEN 
		TIMER(IN := FALSE);
		IO.xPistonOn := FALSE;
		state := 40;
	END_IF
	
	40: // Restart conveyor belts
	NVL_STOPPERING_SEND.isDone := TRUE;
	WaitTime := STRING_TO_TIME('T#1000ms');
	TIMER(IN := TRUE, PT := WaitTime);
	IF TIMER.Q = TRUE THEN 
		TIMER(IN := FALSE);
		state := 15;
	END_IF
	
END_CASE

TIMER();

END_PROGRAM

// Programs/Tools/ErrorFifo
FUNCTION_BLOCK ErrorFifo
VAR_INPUT
	///Input for writing into fifo
	xWrite: BOOL;
	///Input for delete from fifo
	xDelete: BOOL;
	///The error ID
	sErrorID: STRING;
END_VAR
VAR
	///Array for the error table	
	astErrorEvent: ARRAY[1..20] OF st_ErrorEvent;
	///Triger for the rising edge of writing
	rtWrite: R_TRIG;
	///Triger for the rising edge of deleting
	rtDelete: R_TRIG;
	///Variable for the FOR loop
	uiI: UINT;
	///
	dtDateTime: DATE_AND_TIME;
	///Ask the systemtime
	fbGetTime: RTCLK.GetDateAndTime;
	///Variable to store the time data
	sDate: STRING;
	sFormat: STRING;
	rtGetTime: R_TRIG;
	xWriteTrig : BOOL;
	rtGetTimeDone: R_TRIG;
END_VAR
VAR CONSTANT
	///Not used in ARRAY SIZE !!!
	cuiSize: UINT := 20;
END_VAR

